REGION Network 3
   RUNG wire#powerrail
      Mul(in1 := #"HMI.FVR", in2 := #Config.Limits.LL, out => #"MATH.LL")
      { S7_Templates := "[SrcType := Real, DestType := DInt]" } Convert(in := #"MATH.LL", out => #"FVR.LL")
   END_RUNG
   // the same network as SCL:
   #"MATH.LL" := #"HMI.FVR" * #Config.Limits.LL;
   #"FVR.LL" := REAL_TO_DINT(#"MATH.LL");
END_REGION

REGION Network 4
   RUNG wire#powerrail
      Mul(in1 := #"HMI.FVR", in2 := #Config.Limits.L, out => #"MATH.L")
      { S7_Templates := "[SrcType := Real, DestType := DInt]" } Convert(in := #"MATH.L", out => #"FVR.L")
   END_RUNG
   // the same network as SCL:
   #"MATH.L" := #"HMI.FVR" * #Config.Limits.L;
   #"FVR.L" := REAL_TO_DINT(#"MATH.L");
END_REGION

REGION Network 5
   RUNG wire#powerrail
      Mul(in1 := #"HMI.FVR", in2 := #HPR, out => #"MATH.HR")
      { S7_Templates := "[SrcType := Real, DestType := DInt]" } Convert(in := #"MATH.HR", out => #"FVR.HPR")
   END_RUNG
   // the same network as SCL:
   #"MATH.HR" := #"HMI.FVR" * #HPR;
   #"FVR.HPR" := REAL_TO_DINT(#"MATH.HR");
END_REGION

REGION Network 6
   RUNG wire#powerrail
      Mul(in1 := #"HMI.FVR", in2 := #LPR, out => #"MATH.LR")
      { S7_Templates := "[SrcType := Real, DestType := DInt]" } Convert(in := #"MATH.LR", out => #"FVR.LPR")
   END_RUNG
   // the same network as SCL:
   #"MATH.LR" := #"HMI.FVR" * #LPR;
   #"FVR.LPR" := REAL_TO_DINT(#"MATH.LR");
END_REGION

REGION Network 7
   RUNG wire#powerrail
      Mul(in1 := #"HMI.FVR", in2 := #Config.H, out => #"MATH.CONFIG.H")
      { S7_Templates := "[SrcType := Real, DestType := DInt]" } Convert(in := #"MATH.CONFIG.H", out => #"FVR.CONFIG.H")
   END_RUNG
   // the same network as SCL:
   #"MATH.CONFIG.H" := #"HMI.FVR" * #Config.H;
   #"FVR.CONFIG.H" := REAL_TO_DINT(#"MATH.CONFIG.H");
END_REGION

REGION Network 8: Value 1
   RUNG wire#powerrail
      Contact( #V1GA )
      Coil( #V1GA_1 )
   END_RUNG
   // the same network as SCL:
   #V1GA_1 := #V1GA;
END_REGION

REGION Network 9: Value 1
   RUNG wire#powerrail
      Contact( #V2GA )
      Coil( #V2GA_1 )
   END_RUNG
   // the same network as SCL:
   #V2GA_1 := #V2GA;
END_REGION

REGION Network 10: Value 1
   RUNG wire#powerrail
      Contact( #V3GA )
      Coil( #V3GA_1 )
   END_RUNG
   // the same network as SCL:
   #V3GA_1 := #V3GA;
END_REGION

REGION Network 11: Value 1
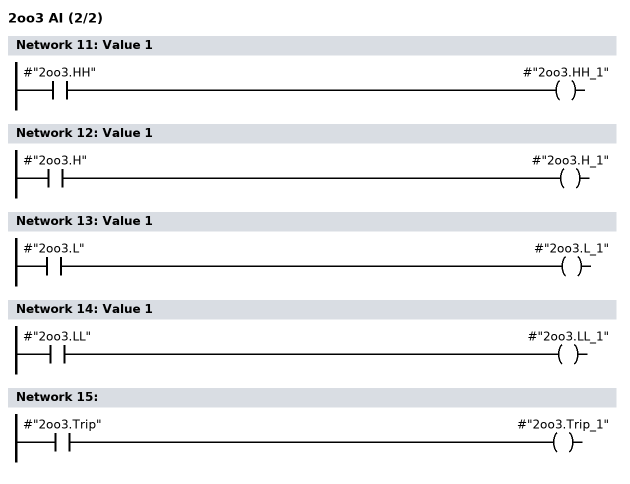
   RUNG wire#powerrail
      Contact( #"2oo3.HH" )
      Coil( #"2oo3.HH_1" )
   END_RUNG
   // the same network as SCL:
   #"2oo3.HH_1" := #"2oo3.HH";
END_REGION

REGION Network 12: Value 1
   RUNG wire#powerrail
      Contact( #"2oo3.H" )
      Coil( #"2oo3.H_1" )
   END_RUNG
   // the same network as SCL:
   #"2oo3.H_1" := #"2oo3.H";
END_REGION

REGION Network 13: Value 1
   RUNG wire#powerrail
      Contact( #"2oo3.L" )
      Coil( #"2oo3.L_1" )
   END_RUNG
   // the same network as SCL:
   #"2oo3.L_1" := #"2oo3.L";
END_REGION

REGION Network 14: Value 1
   RUNG wire#powerrail
      Contact( #"2oo3.LL" )
      Coil( #"2oo3.LL_1" )
   END_RUNG
   // the same network as SCL:
   #"2oo3.LL_1" := #"2oo3.LL";
END_REGION

REGION Network 15
   RUNG wire#powerrail
      Contact( #"2oo3.Trip" )
      Coil( #"2oo3.Trip_1" )
   END_RUNG
   // the same network as SCL:
   #"2oo3.Trip_1" := #"2oo3.Trip";
END_REGION
END_FUNCTION_BLOCK

// folder: 1}Library/Digital

FUNCTION_BLOCK "Signal"   // FB816, LAD
{ S7_Optimized_Access := 'TRUE' }
VERSION : 1.1
   VAR_INPUT
      Mode : Int;   // FB Mode - "0=Interlock N/A" "1=Interlock Used"
      IN : Bool;   // Signal Input
      P : Bool;   // Permissive
      Invert : Bool;   // Invert Output
   END_VAR
   VAR_OUTPUT
      Q : Bool;   // Output
   END_VAR
   VAR_IN_OUT
      REI : Bool;   // Reintegrate
   END_VAR
   VAR
      DBNC_TMR : TON_TIME;
      HLD_TMR : TOF_TIME;
      HMI : Struct
         Controls : Struct
            Pass : Bool;   // Passivate Signal
         END_STRUCT;
         Config : Struct
            DBNC_PT : Time := T#1S;   // Debounce Preset Time
            HLD_PT : Time := T#1S;   // Hold Preset Time
         END_STRUCT;
         Status : Struct
            P : Bool;   // Permissive Status
         END_STRUCT;
      END_STRUCT;
      Reintegrate : "Reintegrate";
   END_VAR
   VAR_TEMP
      ON : Bool;
   END_VAR
BEGIN

REGION Network 1
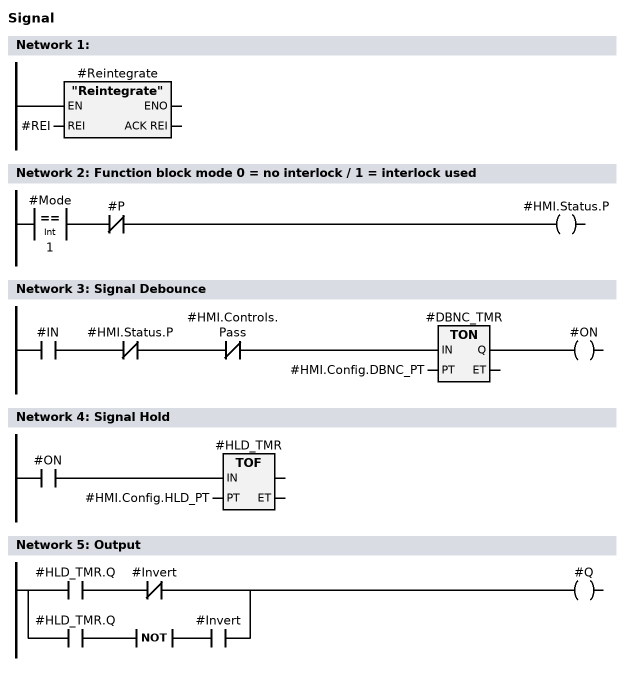
   RUNG wire#powerrail
      #Reintegrate(REI := #REI, "ACK REI" =>)
   END_RUNG
   // the same network as SCL:
   #Reintegrate(REI := #REI);   // "Reintegrate"
END_REGION

REGION Network 2: Function block mode 0 = no interlock / 1 = interlock used
   RUNG wire#powerrail
      { S7_Templates := "SrcType := Int" } EQ_Contact(in1 := #Mode, in2 := 1)
      I_Contact( #P )
      Coil( #HMI.Status.P )
   END_RUNG
   // the same network as SCL:
   #HMI.Status.P := (#Mode = 1) AND NOT #P;
END_REGION

REGION Network 3: Signal Debounce
   #DBNC_TMR(IN := #IN AND NOT #HMI.Status.P AND NOT #HMI.Controls.Pass, PT := #HMI.Config.DBNC_PT);   // TON
   #ON := #DBNC_TMR.Q;
END_REGION

REGION Network 4: Signal Hold
   #HLD_TMR(IN := #ON, PT := #HMI.Config.HLD_PT);   // TOF
END_REGION

REGION Network 5: Output
   RUNG wire#powerrail
      Contact( #HLD_TMR.Q )
      I_Contact( #Invert )
      wire#w1
      Coil( #Q )
   END_RUNG
   RUNG wire#powerrail
      Contact( #HLD_TMR.Q )
      Not()
      Contact( #Invert )
   END_RUNG wire#w1
   // the same network as SCL:
   #Q := (#HLD_TMR.Q AND NOT #Invert) OR (NOT #HLD_TMR.Q AND #Invert);
END_REGION
END_FUNCTION_BLOCK

// folder: 1}Library/E-Stop

FUNCTION_BLOCK "E-STOP"   // FB8, LAD
{ S7_Optimized_Access := 'TRUE' }
VERSION : 0.1
   VAR_INPUT
      ESD1 : Bool := TRUE;
      ESD2 : Bool := TRUE;
      ESD3 : Bool := TRUE;
      ESD4 : Bool := TRUE;
      ESD5 : Bool := TRUE;
      ESD6 : Bool := TRUE;
      ESD7 : Bool := TRUE;
      ESD8 : Bool := TRUE;
      ESD9 : Bool := TRUE;
      ESD10 : Bool := TRUE;
      ESD11 : Bool := TRUE;
      ESD12 : Bool := TRUE;
      ESD13 : Bool := TRUE;
      ESD14 : Bool := TRUE;
      ESD15 : Bool := TRUE;
      ESDD16 : Bool := TRUE;
   END_VAR
   VAR_OUTPUT
      esdActive : Bool;
   END_VAR
   VAR
      masterESD : Bool := TRUE;
      hmiEsd : Bool := TRUE;
      ESDreset : Bool;
   END_VAR
BEGIN

REGION Network 1
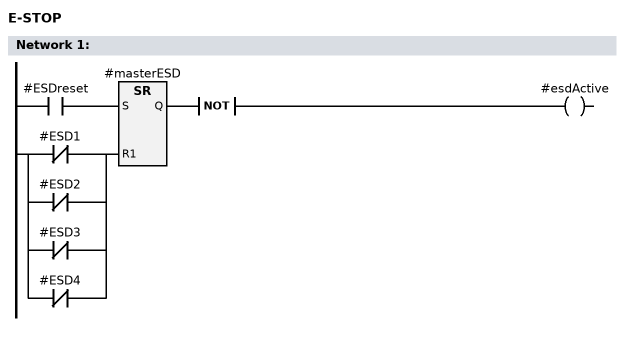
   RUNG wire#powerrail
      Contact( #ESDreset )
      S_SR(operand := #masterESD, r1 := wire#w1)
      Not()
      Coil( #esdActive )
   END_RUNG
   RUNG wire#powerrail
      I_Contact( #ESD1 )
   END_RUNG wire#w1
   RUNG wire#powerrail
      I_Contact( #ESD2 )
   END_RUNG wire#w1
   RUNG wire#powerrail
      I_Contact( #ESD3 )
   END_RUNG wire#w1
   RUNG wire#powerrail
      I_Contact( #ESD4 )
   END_RUNG wire#w1
   // the same network as SCL:
   IF #ESDreset THEN
       #masterESD := TRUE;   // SR flip-flop
   END_IF;
   IF NOT #ESD1 OR NOT #ESD2 OR NOT #ESD3 OR NOT #ESD4 THEN #masterESD := FALSE; END_IF;
   #esdActive := NOT #masterESD;
END_REGION
END_FUNCTION_BLOCK

// folder: 1}Library/Helpers

FUNCTION_BLOCK "Reintegrate"   // FB6, LAD
{ S7_Optimized_Access := 'TRUE' }
VERSION : 0.1
   VAR_OUTPUT
      "ACK REI" : Int;   // Acknowledge Reintegration
   END_VAR
   VAR_IN_OUT
      REI : Bool;   // Reintegrate
   END_VAR
   VAR
      Reintegrating : Bool;
      PT : Struct   // Preset Time
         S1T : Time := T#2s;
         S2T : Time := T#2s;
      END_STRUCT;
      Pulse : Struct
         REI : Bool;
         S1 : Bool;
         S2 : Bool;
         "S2 Q" : Bool;
         Reset : Bool;
      END_STRUCT;
      S1T : TON_TIME;   // Step 1 Timer
      S2T : TOF_TIME;   // Step 2 Timer
   END_VAR
   VAR_TEMP   // added for the SCL form of the ladder/FBD networks
      _w1 : Bool;
      _w2 : Bool;
      _w3 : Bool;
   END_VAR
BEGIN

REGION Network 1
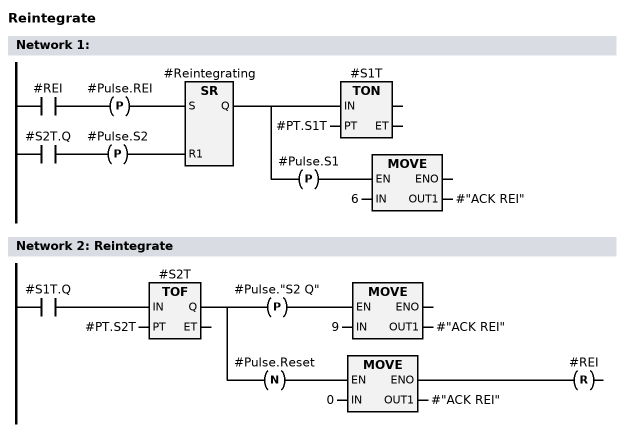
   #_w1 := #REI AND NOT #Pulse.REI;   // rising edge
   #Pulse.REI := #REI;
   #_w2 := #S2T.Q AND NOT #Pulse.S2;   // rising edge
   #Pulse.S2 := #S2T.Q;
   IF #_w1 THEN
       #Reintegrating := TRUE;   // SR flip-flop
   END_IF;
   IF #_w2 THEN #Reintegrating := FALSE; END_IF;
   #S1T(IN := #Reintegrating, PT := #PT.S1T);   // TON
   #_w3 := #Reintegrating AND NOT #Pulse.S1;   // rising edge
   #Pulse.S1 := #Reintegrating;
   IF #_w3 THEN #"ACK REI" := 6; END_IF;
END_REGION

REGION Network 2: Reintegrate
   #S2T(IN := #S1T.Q, PT := #PT.S2T);   // TOF
   #_w1 := #S2T.Q AND NOT #Pulse."S2 Q";   // rising edge
   #Pulse."S2 Q" := #S2T.Q;
   IF #_w1 THEN #"ACK REI" := 9; END_IF;
   #_w2 := NOT #S2T.Q AND #Pulse.Reset;   // falling edge
   #Pulse.Reset := #S2T.Q;
   IF #_w2 THEN
       #"ACK REI" := 0;
       #REI := FALSE;
   END_IF;
END_REGION
END_FUNCTION_BLOCK

FUNCTION_BLOCK "Deviation"   // FB602, LAD
{ S7_Optimized_Access := 'TRUE' }
VERSION : 0.1
   VAR_INPUT
      V1 : Real;   // Value 1 Typically SP
      V2 : Real;   // Value 2 Typically PV
      MXSUV : Real := 1.0;   // Max Step Up Value
      MXSDV : Real := 1.0;   // Max Step Down Value
      MNSUV : Real;   // Min Step Up Value
      MNSDV : Real;   // Min Step Down Value
      UDW : Real := 0.5;   // Upper Deadband Width
      LDW : Real := 0.5;   // Lower Deadband Width
   END_VAR
   VAR_OUTPUT
      DAV : Real;   // Difference Absolute Value
      SU : Bool;   // Step Up = V1 Greater than V2
      SD : Bool;   // Step Down = V1 Less than V2
      V1EQV2 : Bool;   // V1 Equal to V2
      VGTSV : Bool;   // Value Greater Than Step Value
      SUV : Real;   // Step Up Value
      SDV : Real;   // Step Down Value
      DA : Bool;   // Deadband Active
   END_VAR
   VAR
      Status : Struct
         DA : Bool;
         SU : Bool;
         SD : Bool;
         DAV : Real;
      END_STRUCT;
      Deadband : Struct
         UV : Real;   // Upper Value
         LV : Real;   // Lower Value
      END_STRUCT;
   END_VAR
   VAR_TEMP
      N1 : Real;   // V1 - V2
      NMXSDV : Real;   // Negative Max Step Down Value
      TDAV : Real;   // Temp DAV
   END_VAR
BEGIN

REGION Network 1: N1 = |V1 - V2|
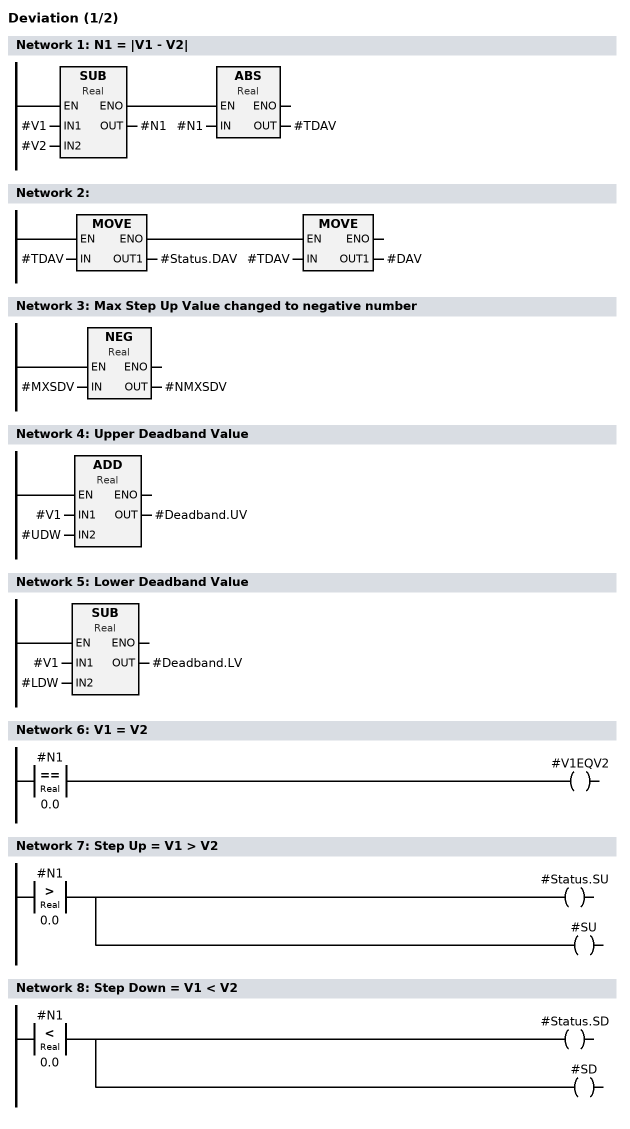
   RUNG wire#powerrail
      { S7_Templates := "SrcType := Real"; S7_GenerateENO := "TRUE" } Sub(in1 := #V1, in2 := #V2, out => #N1)
      { S7_Templates := "SrcType := Real"; S7_GenerateENO := "TRUE" } Abs(in := #N1, out => #TDAV)
   END_RUNG
   // the same network as SCL:
   // ENO of a box is taken as its EN; it also drops when the box reports an error
   #N1 := #V1 - #V2;
   #TDAV := ABS(#N1);
END_REGION

REGION Network 2
   RUNG wire#powerrail
      { S7_GenerateENO := "TRUE" } Move(in := #TDAV, out1 => #Status.DAV)
      { S7_GenerateENO := "TRUE" } Move(in := #TDAV, out1 => #DAV)
   END_RUNG
   // the same network as SCL:
   // ENO of a box is taken as its EN; it also drops when the box reports an error
   #Status.DAV := #TDAV;
   #DAV := #TDAV;
END_REGION

REGION Network 3: Max Step Up Value changed to negative number
   RUNG wire#powerrail
      { S7_Templates := "SrcType := Real"; S7_GenerateENO := "TRUE" } Neg(in := #MXSDV, out => #NMXSDV)
   END_RUNG
   // the same network as SCL:
   #NMXSDV := -#MXSDV;
END_REGION

REGION Network 4: Upper Deadband Value
   RUNG wire#powerrail
      { S7_Templates := "SrcType := Real"; S7_GenerateENO := "TRUE" } Add(in1 := #V1, in2 := #UDW, out => #Deadband.UV)
   END_RUNG
   // the same network as SCL:
   #Deadband.UV := #V1 + #UDW;
END_REGION

REGION Network 5: Lower Deadband Value
   RUNG wire#powerrail
      { S7_Templates := "SrcType := Real"; S7_GenerateENO := "TRUE" } Sub(in1 := #V1, in2 := #LDW, out => #Deadband.LV)
   END_RUNG
   // the same network as SCL:
   #Deadband.LV := #V1 - #LDW;
END_REGION

REGION Network 6: V1 = V2
   RUNG wire#powerrail
      { S7_Templates := "SrcType := Real" } EQ_Contact(in1 := #N1, in2 := 0.0)
      Coil( #V1EQV2 )
   END_RUNG
   // the same network as SCL:
   #V1EQV2 := #N1 = 0.0;
END_REGION

REGION Network 7: Step Up = V1 > V2
   RUNG wire#powerrail
      { S7_Templates := "SrcType := Real" } GT_Contact(in1 := #N1, in2 := 0.0)
      wire#w1
      Coil( #Status.SU )
   END_RUNG
   RUNG wire#w1
      Coil( #SU )
   END_RUNG
   // the same network as SCL:
   #Status.SU := #N1 > 0.0;
   #SU := #Status.SU;
END_REGION

REGION Network 8: Step Down = V1 < V2
   RUNG wire#powerrail
      { S7_Templates := "SrcType := Real" } LT_Contact(in1 := #N1, in2 := 0.0)
      wire#w1
      Coil( #Status.SD )
   END_RUNG
   RUNG wire#w1
      Coil( #SD )
   END_RUNG
   // the same network as SCL:
   #Status.SD := #N1 < 0.0;
   #SD := #Status.SD;
END_REGION

REGION Network 9: Step Up Reached
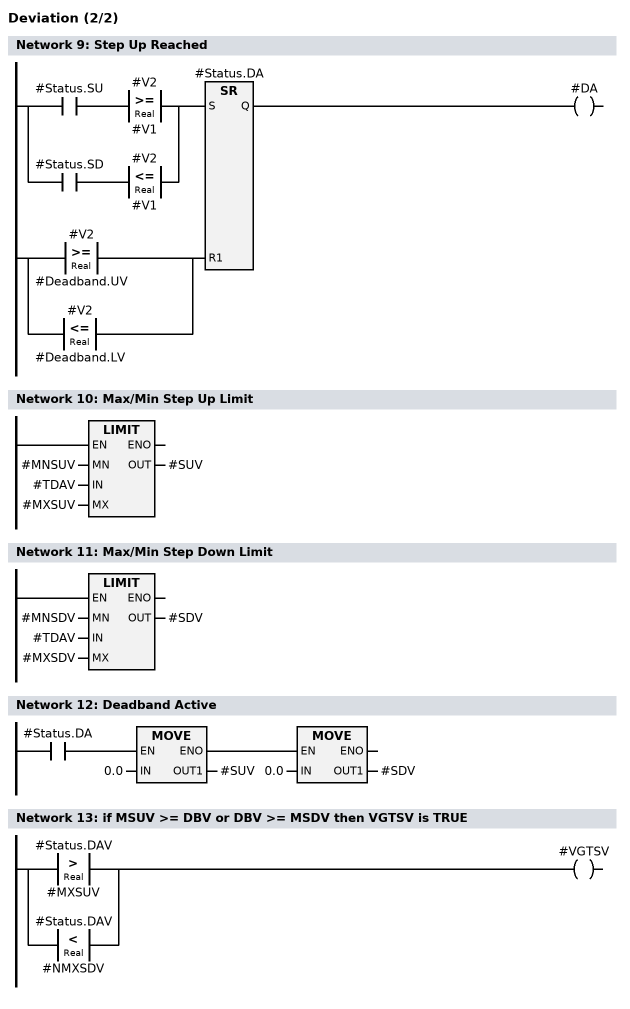
   RUNG wire#powerrail
      Contact( #Status.SU )
      { S7_Templates := "SrcType := Real" } GE_Contact(in1 := #V2, in2 := #V1)
      wire#w1
      S_SR(operand := #Status.DA, r1 := wire#w2)
      Coil( #DA )
   END_RUNG
   RUNG wire#powerrail
      Contact( #Status.SD )
      { S7_Templates := "SrcType := Real" } LE_Contact(in1 := #V2, in2 := #V1)
   END_RUNG wire#w1
   RUNG wire#powerrail
      { S7_Templates := "SrcType := Real" } GE_Contact(in1 := #V2, in2 := #Deadband.UV)
   END_RUNG wire#w2
   RUNG wire#powerrail
      { S7_Templates := "SrcType := Real" } LE_Contact(in1 := #V2, in2 := #Deadband.LV)
   END_RUNG wire#w2
   // the same network as SCL:
   IF (#Status.SU AND (#V2 >= #V1)) OR (#Status.SD AND (#V2 <= #V1)) THEN
       #Status.DA := TRUE;   // SR flip-flop
   END_IF;
   IF (#V2 >= #Deadband.UV) OR (#V2 <= #Deadband.LV) THEN #Status.DA := FALSE; END_IF;
   #DA := #Status.DA;
END_REGION

REGION Network 10: Max/Min Step Up Limit
   #SUV := LIMIT(MN := #MNSUV, IN := #TDAV, MX := #MXSUV);
END_REGION

REGION Network 11: Max/Min Step Down Limit
   #SDV := LIMIT(MN := #MNSDV, IN := #TDAV, MX := #MXSDV);
END_REGION

REGION Network 12: Deadband Active
   RUNG wire#powerrail
      Contact( #Status.DA )
      { S7_GenerateENO := "TRUE" } Move(in := 0.0, out1 => #SUV)
      { S7_GenerateENO := "TRUE" } Move(in := 0.0, out1 => #SDV)
   END_RUNG
   // the same network as SCL:
   // ENO of a box is taken as its EN; it also drops when the box reports an error
   IF #Status.DA THEN
       #SUV := 0.0;
       #SDV := 0.0;
   END_IF;
END_REGION

REGION Network 13: if MSUV >= DBV or DBV >= MSDV then VGTSV is TRUE
   RUNG wire#powerrail
      { S7_Templates := "SrcType := Real" } GT_Contact(in1 := #Status.DAV, in2 := #MXSUV)
      wire#w1
      Coil( #VGTSV )
   END_RUNG
   RUNG wire#powerrail
      { S7_Templates := "SrcType := Real" } LT_Contact(in1 := #Status.DAV, in2 := #NMXSDV)
   END_RUNG wire#w1
   // the same network as SCL:
   #VGTSV := (#Status.DAV > #MXSUV) OR (#Status.DAV < #NMXSDV);
END_REGION
END_FUNCTION_BLOCK

FUNCTION_BLOCK "HLR"   // FB720, LAD
TITLE = High Limit REAL
{ S7_Optimized_Access := 'TRUE' }
VERSION : 0.3
   VAR_INPUT
      IV : Real;   // Input Value
      HL : Real;   // High Limit
      H : Real;   // Hysteresis
      PM : Int;   // Permissive Mode - "0=No P""1=Bool P" "2=Real P"
      PB : Bool;   // Permissive BOOL
      PR : Real;   // Permissive REAL
   END_VAR
   VAR_OUTPUT
      LR : Bool;   // Limit Reached
   END_VAR
   VAR
      Config : Struct
         DPT : Time := T#1S;   // Debounce Preset Time
         HPT : Time := T#1S;   // Hold Preset Time
         PPT : Time := T#10S;   // Permissive Preset Time
         PSP : Real;   // Permissive Setpoint
         PRS : Real;   // Permissive Reset Setpoint
      END_STRUCT;
      Admin : Struct
         HV : Real;   // Hysteresis Value
         SL : Bool;   // SR Limit
         PA : Bool;   // Permissive Active
         AR : Bool;   // Alarm Reset (Only used during a mode change)
      END_STRUCT;
      DBT : TON_TIME;   // Debounce Timer
      HT : TOF_TIME;   // Hold Timer
      PT : TON_TIME;   // Permissive Class B Timer
   END_VAR
   VAR_TEMP   // added for the SCL form of the ladder/FBD networks
      _w1 : Bool;
      _w2 : Bool;
   END_VAR
BEGIN

REGION Network 1: Permissive Mode 2 Logic
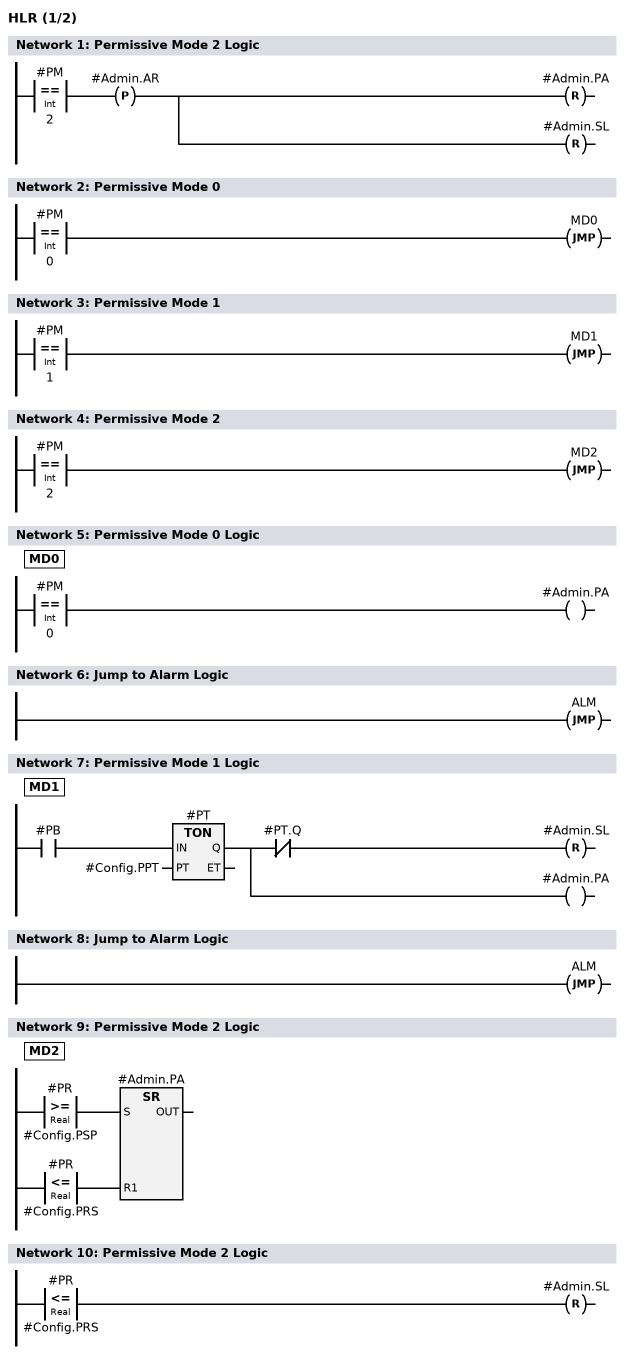
   RUNG wire#powerrail
      { S7_Templates := "SrcType := Int" } EQ_Contact(in1 := #PM, in2 := 2)
      P_Trig( #Admin.AR )
      wire#w1
      R_Coil( #Admin.PA )
   END_RUNG
   RUNG wire#w1
      R_Coil( #Admin.SL )
   END_RUNG
   // the same network as SCL:
   #_w1 := #PM = 2;
   #_w2 := #_w1 AND NOT #Admin.AR;   // rising edge
   #Admin.AR := #_w1;
   IF #_w2 THEN
       #Admin.PA := FALSE;
       #Admin.SL := FALSE;
   END_IF;
END_REGION

REGION Network 2: Permissive Mode 0
   RUNG wire#powerrail
      { S7_Templates := "SrcType := Int" } EQ_Contact(in1 := #PM, in2 := 0)
      JumpCoil( MD0 )
   END_RUNG
   // the same network as SCL:
   IF #PM = 0 THEN GOTO MD0; END_IF;
END_REGION

REGION Network 3: Permissive Mode 1
   RUNG wire#powerrail
      { S7_Templates := "SrcType := Int" } EQ_Contact(in1 := #PM, in2 := 1)
      JumpCoil( MD1 )
   END_RUNG
   // the same network as SCL:
   IF #PM = 1 THEN GOTO MD1; END_IF;
END_REGION

REGION Network 4: Permissive Mode 2
   RUNG wire#powerrail
      { S7_Templates := "SrcType := Int" } EQ_Contact(in1 := #PM, in2 := 2)
      JumpCoil( MD2 )
   END_RUNG
   // the same network as SCL:
   IF #PM = 2 THEN GOTO MD2; END_IF;
END_REGION

REGION Network 5: Permissive Mode 0 Logic
   Label( MD0 )
   RUNG wire#powerrail
      { S7_Templates := "SrcType := Int" } EQ_Contact(in1 := #PM, in2 := 0)
      Coil( #Admin.PA )
   END_RUNG
   // the same network as SCL:
   MD0:
   #Admin.PA := #PM = 0;
END_REGION

REGION Network 6: Jump to Alarm Logic
   RUNG wire#powerrail
      JumpCoil( ALM )
   END_RUNG
   // the same network as SCL:
   GOTO ALM;
END_REGION

REGION Network 7: Permissive Mode 1 Logic
   MD1:
   #PT(IN := #PB, PT := #Config.PPT);   // TON
   IF #PT.Q AND NOT #PT.Q THEN #Admin.SL := FALSE; END_IF;
   #Admin.PA := #PT.Q;
END_REGION

REGION Network 8: Jump to Alarm Logic
   RUNG wire#powerrail
      JumpCoil( ALM )
   END_RUNG
   // the same network as SCL:
   GOTO ALM;
END_REGION

REGION Network 9: Permissive Mode 2 Logic
   Label( MD2 )
   RUNG wire#powerrail
      { S7_Templates := "SrcType := Real" } GE_Contact(in1 := #PR, in2 := #Config.PSP)
      S_SR(operand := #Admin.PA, r1 := wire#w1)
   END_RUNG
   RUNG wire#powerrail
      { S7_Templates := "SrcType := Real" } LE_Contact(in1 := #PR, in2 := #Config.PRS)
   END_RUNG wire#w1
   // the same network as SCL:
   MD2:
   IF #PR >= #Config.PSP THEN
       #Admin.PA := TRUE;   // SR flip-flop
   END_IF;
   IF #PR <= #Config.PRS THEN #Admin.PA := FALSE; END_IF;
END_REGION

REGION Network 10: Permissive Mode 2 Logic
   RUNG wire#powerrail
      { S7_Templates := "SrcType := Real" } LE_Contact(in1 := #PR, in2 := #Config.PRS)
      R_Coil( #Admin.SL )
   END_RUNG
   // the same network as SCL:
   IF #PR <= #Config.PRS THEN #Admin.SL := FALSE; END_IF;
END_REGION

REGION Network 11: Jump to Alarm Logic
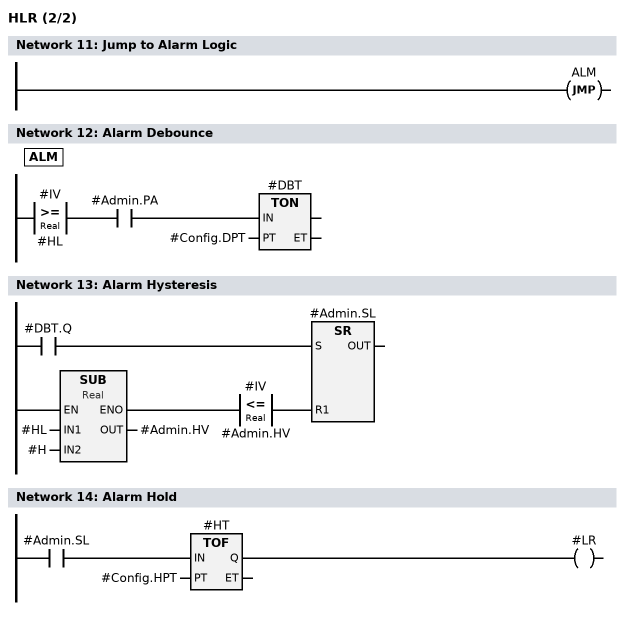
   RUNG wire#powerrail
      JumpCoil( ALM )
   END_RUNG
   // the same network as SCL:
   GOTO ALM;
END_REGION

REGION Network 12: Alarm Debounce
   ALM:
   #DBT(IN := (#IV >= #HL) AND #Admin.PA, PT := #Config.DPT);   // TON
END_REGION

REGION Network 13: Alarm Hysteresis
   RUNG wire#powerrail
      Contact( #DBT.Q )
      S_SR(operand := #Admin.SL, r1 := wire#w1)
   END_RUNG
   RUNG wire#powerrail
      { S7_Templates := "SrcType := Real"; S7_GenerateENO := "TRUE" } Sub(in1 := #HL, in2 := #H, out => #Admin.HV)
      { S7_Templates := "SrcType := Real" } LE_Contact(in1 := #IV, in2 := #Admin.HV)
   END_RUNG wire#w1
   // the same network as SCL:
   // ENO of a box is taken as its EN; it also drops when the box reports an error
   #Admin.HV := #HL - #H;
   IF #DBT.Q THEN
       #Admin.SL := TRUE;   // SR flip-flop
   END_IF;
   IF #IV <= #Admin.HV THEN #Admin.SL := FALSE; END_IF;
END_REGION

REGION Network 14: Alarm Hold
   #HT(IN := #Admin.SL, PT := #Config.HPT);   // TOF
   #LR := #HT.Q;
END_REGION
END_FUNCTION_BLOCK

FUNCTION_BLOCK "LLR"   // FB721, LAD
TITLE = Low Limit REAL
{ S7_Optimized_Access := 'TRUE' }
VERSION : 0.2
   VAR_INPUT
      IV : Real;   // Input Value
      LL : Real;   // Low Limit
      H : Real;   // Hysteresis
      PM : Int;   // Permissive Mode - "0=No P""1=Bool P" "2=Real P"
      PB : Bool;   // Permissive BOOL
      PR : Real;   // Permissive REAL
   END_VAR
   VAR_OUTPUT
      LR : Bool;   // Limit Reached
   END_VAR
   VAR
      Config : Struct
         DPT : Time := T#1S;   // Debounce Preset Time
         HPT : Time := T#1S;   // Hold Preset Time
         PPT : Time := T#10S;   // Permissive Preset Time
         PSP : Real;   // Permissive Setpoint
         PRS : Real;   // Permissive Reset Setpoint
      END_STRUCT;
      Admin : Struct
         HV : Real;   // Hysteresis Value
         SL : Bool;   // SR Limit
         PA : Bool;   // Permissive Active
         AR : Bool;   // Alarm Reset (Only used during a mode change)
      END_STRUCT;
      DBT : TON_TIME;   // Debounce Timer
      HT : TOF_TIME;   // Hold Timer
      PT : TON_TIME;   // Permissive Class B Timer
   END_VAR
   VAR_TEMP   // added for the SCL form of the ladder/FBD networks
      _w1 : Bool;
      _w2 : Bool;
   END_VAR
BEGIN

REGION Network 1: Permissive Mode 2 Logic
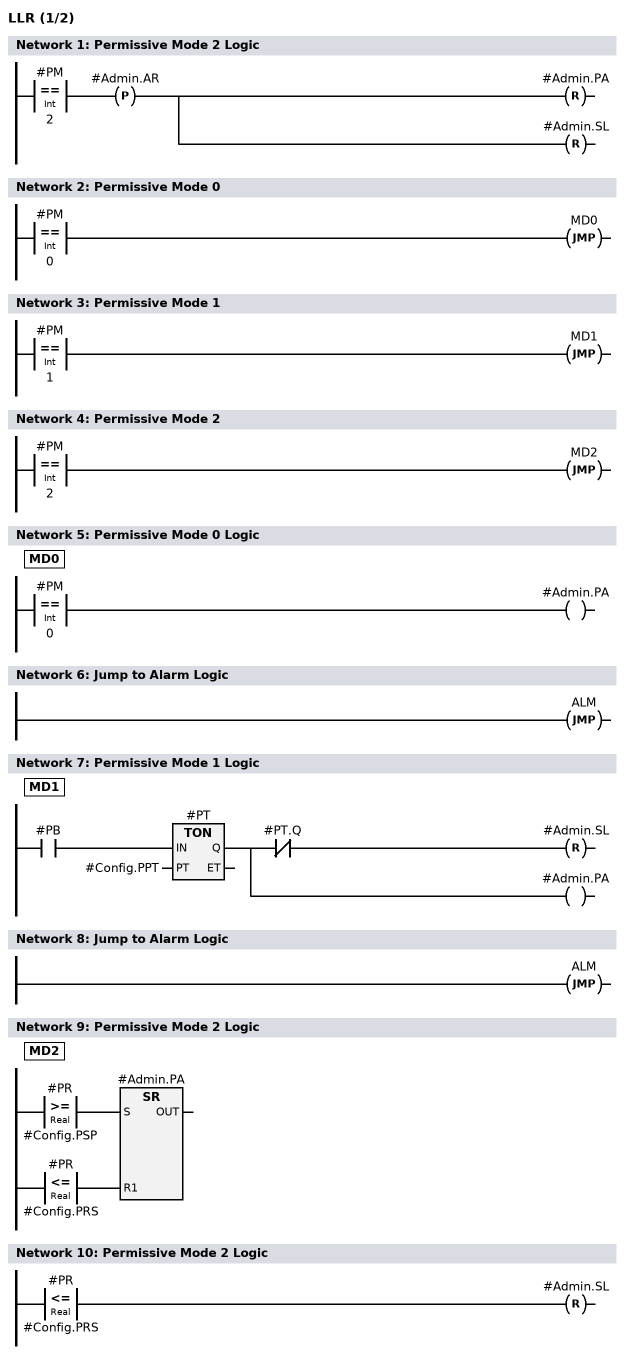
   RUNG wire#powerrail
      { S7_Templates := "SrcType := Int" } EQ_Contact(in1 := #PM, in2 := 2)
      P_Trig( #Admin.AR )
      wire#w1
      R_Coil( #Admin.PA )
   END_RUNG
   RUNG wire#w1
      R_Coil( #Admin.SL )
   END_RUNG
   // the same network as SCL:
   #_w1 := #PM = 2;
   #_w2 := #_w1 AND NOT #Admin.AR;   // rising edge
   #Admin.AR := #_w1;
   IF #_w2 THEN
       #Admin.PA := FALSE;
       #Admin.SL := FALSE;
   END_IF;
END_REGION

REGION Network 2: Permissive Mode 0
   RUNG wire#powerrail
      { S7_Templates := "SrcType := Int" } EQ_Contact(in1 := #PM, in2 := 0)
      JumpCoil( MD0 )
   END_RUNG
   // the same network as SCL:
   IF #PM = 0 THEN GOTO MD0; END_IF;
END_REGION

REGION Network 3: Permissive Mode 1
   RUNG wire#powerrail
      { S7_Templates := "SrcType := Int" } EQ_Contact(in1 := #PM, in2 := 1)
      JumpCoil( MD1 )
   END_RUNG
   // the same network as SCL:
   IF #PM = 1 THEN GOTO MD1; END_IF;
END_REGION

REGION Network 4: Permissive Mode 2
   RUNG wire#powerrail
      { S7_Templates := "SrcType := Int" } EQ_Contact(in1 := #PM, in2 := 2)
      JumpCoil( MD2 )
   END_RUNG
   // the same network as SCL:
   IF #PM = 2 THEN GOTO MD2; END_IF;
END_REGION

REGION Network 5: Permissive Mode 0 Logic
   Label( MD0 )
   RUNG wire#powerrail
      { S7_Templates := "SrcType := Int" } EQ_Contact(in1 := #PM, in2 := 0)
      Coil( #Admin.PA )
   END_RUNG
   // the same network as SCL:
   MD0:
   #Admin.PA := #PM = 0;
END_REGION

REGION Network 6: Jump to Alarm Logic
   RUNG wire#powerrail
      JumpCoil( ALM )
   END_RUNG
   // the same network as SCL:
   GOTO ALM;
END_REGION

REGION Network 7: Permissive Mode 1 Logic
   MD1:
   #PT(IN := #PB, PT := #Config.PPT);   // TON
   IF #PT.Q AND NOT #PT.Q THEN #Admin.SL := FALSE; END_IF;
   #Admin.PA := #PT.Q;
END_REGION

REGION Network 8: Jump to Alarm Logic
   RUNG wire#powerrail
      JumpCoil( ALM )
   END_RUNG
   // the same network as SCL:
   GOTO ALM;
END_REGION

REGION Network 9: Permissive Mode 2 Logic
   Label( MD2 )
   RUNG wire#powerrail
      { S7_Templates := "SrcType := Real" } GE_Contact(in1 := #PR, in2 := #Config.PSP)
      S_SR(operand := #Admin.PA, r1 := wire#w1)
   END_RUNG
   RUNG wire#powerrail
      { S7_Templates := "SrcType := Real" } LE_Contact(in1 := #PR, in2 := #Config.PRS)
   END_RUNG wire#w1
   // the same network as SCL:
   MD2:
   IF #PR >= #Config.PSP THEN
       #Admin.PA := TRUE;   // SR flip-flop
   END_IF;
   IF #PR <= #Config.PRS THEN #Admin.PA := FALSE; END_IF;
END_REGION

REGION Network 10: Permissive Mode 2 Logic
   RUNG wire#powerrail
      { S7_Templates := "SrcType := Real" } LE_Contact(in1 := #PR, in2 := #Config.PRS)
      R_Coil( #Admin.SL )
   END_RUNG
   // the same network as SCL:
   IF #PR <= #Config.PRS THEN #Admin.SL := FALSE; END_IF;
END_REGION

REGION Network 11: Jump to Alarm Logic
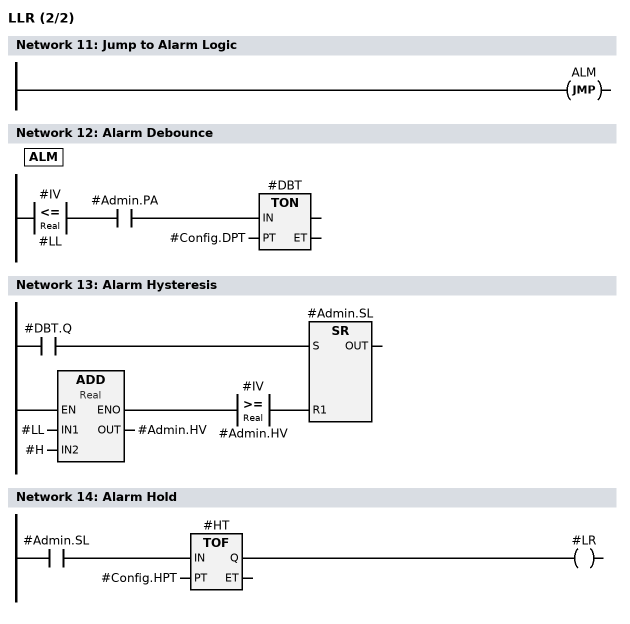
   RUNG wire#powerrail
      JumpCoil( ALM )
   END_RUNG
   // the same network as SCL:
   GOTO ALM;
END_REGION

REGION Network 12: Alarm Debounce
   ALM:
   #DBT(IN := (#IV <= #LL) AND #Admin.PA, PT := #Config.DPT);   // TON
END_REGION

REGION Network 13: Alarm Hysteresis
   RUNG wire#powerrail
      Contact( #DBT.Q )
      S_SR(operand := #Admin.SL, r1 := wire#w1)
   END_RUNG
   RUNG wire#powerrail
      { S7_Templates := "SrcType := Real"; S7_GenerateENO := "TRUE" } Add(in1 := #LL, in2 := #H, out => #Admin.HV)
      { S7_Templates := "SrcType := Real" } GE_Contact(in1 := #IV, in2 := #Admin.HV)
   END_RUNG wire#w1
   // the same network as SCL:
   // ENO of a box is taken as its EN; it also drops when the box reports an error
   #Admin.HV := #LL + #H;
   IF #DBT.Q THEN
       #Admin.SL := TRUE;   // SR flip-flop
   END_IF;
   IF #IV >= #Admin.HV THEN #Admin.SL := FALSE; END_IF;
END_REGION

REGION Network 14: Alarm Hold
   #HT(IN := #Admin.SL, PT := #Config.HPT);   // TOF
   #LR := #HT.Q;
END_REGION
END_FUNCTION_BLOCK

FUNCTION_BLOCK "Max 2R"   // FB722, LAD
{ S7_Optimized_Access := 'TRUE' }
VERSION : 0.1
   VAR_INPUT
      V1 : Real;   // Value 1
      V2 : Real;   // Value 2
   END_VAR
   VAR_OUTPUT
      FV : Real;   // Final Value
      V1A : Bool;   // Value 1 Active
      V2A : Bool;   // Value 2 Active
   END_VAR
   VAR_TEMP   // added for the SCL form of the ladder/FBD networks
      _w1 : Bool;
   END_VAR
BEGIN

REGION Network 1: Value 1 Active
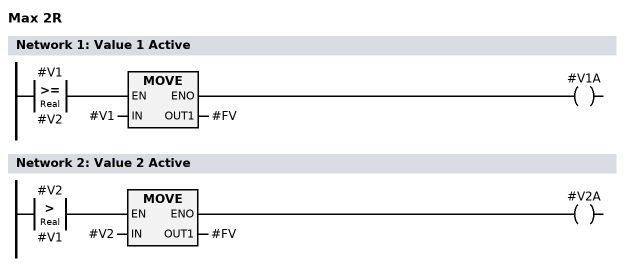
   RUNG wire#powerrail
      { S7_Templates := "SrcType := Real" } GE_Contact(in1 := #V1, in2 := #V2)
      { S7_GenerateENO := "TRUE" } Move(in := #V1, out1 => #FV)
      Coil( #V1A )
   END_RUNG
   // the same network as SCL:
   // ENO of a box is taken as its EN; it also drops when the box reports an error
   #_w1 := #V1 >= #V2;
   IF #_w1 THEN #FV := #V1; END_IF;
   #V1A := #_w1;
END_REGION

REGION Network 2: Value 2 Active
   RUNG wire#powerrail
      { S7_Templates := "SrcType := Real" } GT_Contact(in1 := #V2, in2 := #V1)
      { S7_GenerateENO := "TRUE" } Move(in := #V2, out1 => #FV)
      Coil( #V2A )
   END_RUNG
   // the same network as SCL:
   // ENO of a box is taken as its EN; it also drops when the box reports an error
   #_w1 := #V2 > #V1;
   IF #_w1 THEN #FV := #V2; END_IF;
   #V2A := #_w1;
END_REGION
END_FUNCTION_BLOCK

FUNCTION_BLOCK "Min 2R"   // FB723, LAD
{ S7_Optimized_Access := 'TRUE' }
VERSION : 0.1
   VAR_INPUT
      V1 : Real;   // Value 1
      V2 : Real;   // Value 2
   END_VAR
   VAR_OUTPUT
      FV : Real;   // Final Value
      V1A : Bool;   // Value 1 Active
      V2A : Bool;   // Value 2 Active
   END_VAR
   VAR_TEMP   // added for the SCL form of the ladder/FBD networks
      _w1 : Bool;
   END_VAR
BEGIN

REGION Network 1: Value 1 Active
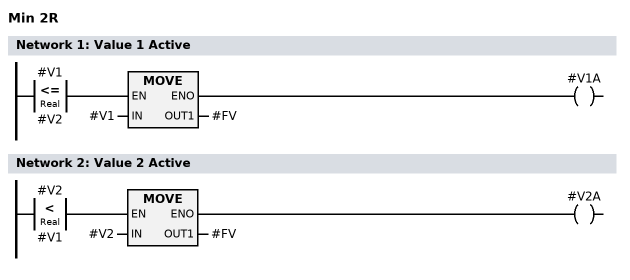
   RUNG wire#powerrail
      { S7_Templates := "SrcType := Real" } LE_Contact(in1 := #V1, in2 := #V2)
      { S7_GenerateENO := "TRUE" } Move(in := #V1, out1 => #FV)
      Coil( #V1A )
   END_RUNG
   // the same network as SCL:
   // ENO of a box is taken as its EN; it also drops when the box reports an error
   #_w1 := #V1 <= #V2;
   IF #_w1 THEN #FV := #V1; END_IF;
   #V1A := #_w1;
END_REGION

REGION Network 2: Value 2 Active
   RUNG wire#powerrail
      { S7_Templates := "SrcType := Real" } LT_Contact(in1 := #V2, in2 := #V1)
      { S7_GenerateENO := "TRUE" } Move(in := #V2, out1 => #FV)
      Coil( #V2A )
   END_RUNG
   // the same network as SCL:
   // ENO of a box is taken as its EN; it also drops when the box reports an error
   #_w1 := #V2 < #V1;
   IF #_w1 THEN #FV := #V2; END_IF;
   #V2A := #_w1;
END_REGION
END_FUNCTION_BLOCK

FUNCTION "USAV" : Void   // FC1, LAD
{ S7_Optimized_Access := 'TRUE' }
VERSION : 0.1
   VAR_INPUT
      Value : Real;   // Final Scaled Analog Input
      EMXV : Real;   // Engineering Max Value
      EMNV : Real;   // Engineering Min Value
      RMXV : Int;   // Raw Max Value
      RMNV : Int;   // Raw Min Value
   END_VAR
   VAR_OUTPUT
      AOI : Int;   // Analog Output INT
   END_VAR
   VAR_TEMP
      AIOV : Real;   // Analog Input Output Value
   END_VAR
BEGIN

REGION Network 1: Normalize and Unscale the value
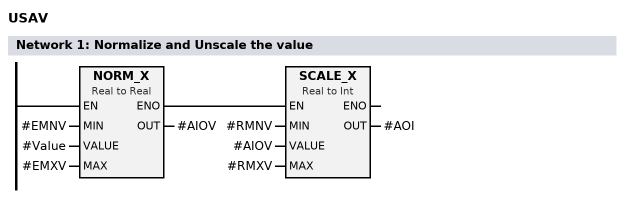
   RUNG wire#powerrail
      { S7_Templates := "[SrcType := Real, DestType := Real]" } Normalize(min := #EMNV, value := #Value, max := #EMXV, out => #AIOV)
      { S7_Templates := "[SrcType := Real, DestType := Int]" } Scale(min := #RMNV, value := #AIOV, max := #RMXV, out => #AOI)
   END_RUNG
   // the same network as SCL:
   #AIOV := NORM_X(MIN := #EMNV, VALUE := #Value, MAX := #EMXV);
   #AOI := SCALE_X(MIN := #RMNV, VALUE := #AIOV, MAX := #RMXV);
END_REGION
END_FUNCTION

FUNCTION "PIDnormMove" : Void   // FC3, LAD
{ S7_Optimized_Access := 'TRUE' }
VERSION : 0.1
   VAR_INPUT
      normalizedEnabled : Bool;
      Emax1 : Real;
      Emin1 : Real;
      Pv1 : Real;
      Emax2 : Real;
      Emin2 : Real;
      Pv2 : Real;
   END_VAR
   VAR_OUTPUT
      Emax : Real;
      Emin : Real;
      PV : Real;
   END_VAR
BEGIN

REGION Network 1
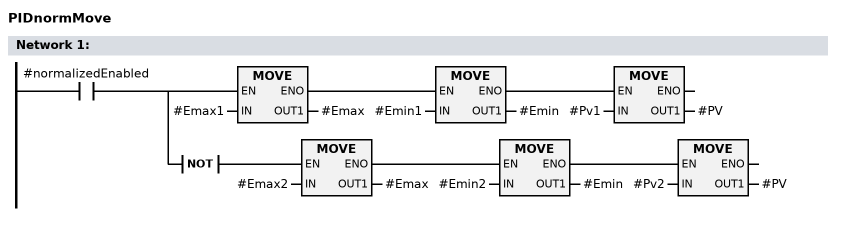
   RUNG wire#powerrail
      Contact( #normalizedEnabled )
      wire#w1
      Move(in := #Emax1, out1 => #Emax)
      Move(in := #Emin1, out1 => #Emin)
      Move(in := #Pv1, out1 => #PV)
   END_RUNG
   RUNG wire#w1
      Not()
      Move(in := #Emax2, out1 => #Emax)
      Move(in := #Emin2, out1 => #Emin)
      Move(in := #Pv2, out1 => #PV)
   END_RUNG
   // the same network as SCL:
   IF #normalizedEnabled THEN
       #Emax := #Emax1;
       #Emin := #Emin1;
       #PV := #Pv1;
   END_IF;
   IF NOT #normalizedEnabled THEN
       #Emax := #Emax2;
       #Emin := #Emin2;
       #PV := #Pv2;
   END_IF;
END_REGION
END_FUNCTION

FUNCTION "Range" : Void   // FC700, LAD
{ S7_Optimized_Access := 'FALSE' }
VERSION : 0.1
   VAR_INPUT
      PV : Real;
      SP : Real;
      UR_DB_SP : Real;   // Upper Range Deadband Setpoint
      LR_DB_SP : Real;   // Lower Range Deadband Setpoint
   END_VAR
   VAR_OUTPUT
      WR : Bool;   // Within Range
      UR_Val : Real;
      LR_Val : Real;
   END_VAR
   VAR_TEMP
      "UR Value" : Real;
      "LR Value" : Real;
   END_VAR
BEGIN

REGION Network 1: Upper & Lower Range
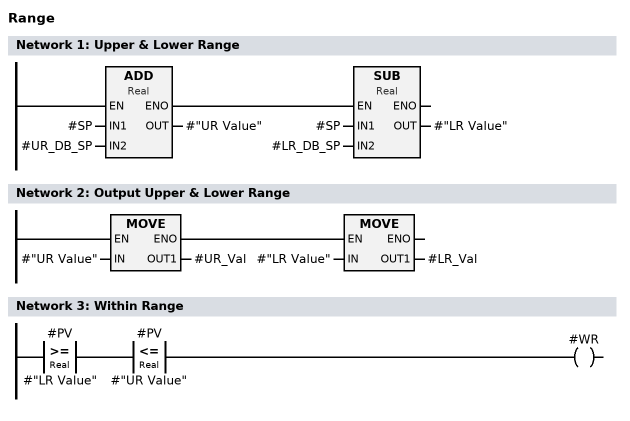
   RUNG wire#powerrail
      { S7_Templates := "SrcType := Real"; S7_GenerateENO := "TRUE" } Add(in1 := #SP, in2 := #UR_DB_SP, out => #"UR Value")
      { S7_Templates := "SrcType := Real"; S7_GenerateENO := "TRUE" } Sub(in1 := #SP, in2 := #LR_DB_SP, out => #"LR Value")
   END_RUNG
   // the same network as SCL:
   // ENO of a box is taken as its EN; it also drops when the box reports an error
   #"UR Value" := #SP + #UR_DB_SP;
   #"LR Value" := #SP - #LR_DB_SP;
END_REGION

REGION Network 2: Output Upper & Lower Range
   RUNG wire#powerrail
      { S7_GenerateENO := "TRUE" } Move(in := #"UR Value", out1 => #UR_Val)
      { S7_GenerateENO := "TRUE" } Move(in := #"LR Value", out1 => #LR_Val)
   END_RUNG
   // the same network as SCL:
   // ENO of a box is taken as its EN; it also drops when the box reports an error
   #UR_Val := #"UR Value";
   #LR_Val := #"LR Value";
END_REGION

REGION Network 3: Within Range
   RUNG wire#powerrail
      { S7_Templates := "SrcType := Real" } GE_Contact(in1 := #PV, in2 := #"LR Value")
      { S7_Templates := "SrcType := Real" } LE_Contact(in1 := #PV, in2 := #"UR Value")
      Coil( #WR )
   END_RUNG
   // the same network as SCL:
   #WR := (#PV >= #"LR Value") AND (#PV <= #"UR Value");
END_REGION
END_FUNCTION

FUNCTION "SAV" : Void   // FC900, LAD
{ S7_Optimized_Access := 'FALSE' }
VERSION : 0.2
   VAR_INPUT
      VALUE : Int;   // Analog Input INT
      EMXV : Real;   // Engineering Max Value
      EMNV : Real;   // Engineering Min Value
      RMXV : Int;   // Raw Max Value
      RMNV : Int;   // Raw Min Value
   END_VAR
   VAR_OUTPUT
      SAI : Real;   // Final Scaled Analog Input
   END_VAR
   VAR_TEMP
      AIOV : Real;   // Analog Input Output Value
   END_VAR
BEGIN

REGION Network 1
